// TIA Portal project "ESTHER_Gas_v4.0_4" (V13)

(* hardware
DEVICE "SIMATIC 1200 station_1"  S71200.Device
   slot 0: "S7-1200 rack"  Rack  V1.0
   slot 1: "PLC_1"  CPU 1215C DC/DC/DC  6ES7 215-1AG40-0XB0  V4.1
   slot 2: "DQ 16x24VDC_1"  6ES7 222-1BH32-0XB0  V2.0
   slot 3: "AI 8x13BIT_1"  6ES7 231-4HF32-0XB0  V2.0
   slot 4: "AI 8x13BIT_2"  6ES7 231-4HF32-0XB0  V2.0
   slot 101: "CM 1241 (RS422/485)_1"  6ES7 241-1CH32-0XB0  V2.1
   slot 102: "CM 1241 (RS422/485)_2"  6ES7 241-1CH32-0XB0  V2.1
*)

// ===== PLC "PLC_1"  CPU 1215C DC/DC/DC =====

VAR_GLOBAL   // PLC tag table "Default tag table"
   "PV701_NOT_CLOSED_LS" AT %I0.0 : Bool;   // PV701 Limit Switch
   "PV701_NOT_OPEN_LS" AT %I0.1 : Bool;   // PV701 Limit Switch
   "PV702_NOT_CLOSED_LS" AT %I0.2 : Bool;   // PV702 Limit Switch
   "PV702_NOT_OPEN_LS" AT %I0.3 : Bool;   // PV702 Limit Switch
   "PV703A_NOT_OPEN_LS" AT %I0.4 : Bool;
   "PV703A_NOT_CLOSED_LS" AT %I0.5 : Bool;
   "PV703B_NOT_OPEN_LS" AT %I0.6 : Bool;
   "PV703B_NOT_CLOSED_LS" AT %I0.7 : Bool;
   "PT101_ADC" AT %IW114 : Word;
   "PV101_NC" AT %Q9.3 : Bool;   // NC
   "PV102_NO" AT %Q9.4 : Bool;   // NO Temp
   "STEP_0_ON" AT %Q1.7 : Bool;
   "STEP_1_ON" AT %Q1.2 : Bool;
   "STEP_2_ON" AT %Q1.3 : Bool;
   "STEP_3_ON" AT %Q1.4 : Bool;
   "PV201_NC" AT %Q8.3 : Bool;
   "PV301_NC" AT %Q8.6 : Bool;
   "PV401_NC" AT %Q8.0 : Bool;
   "PV202_NC" AT %Q8.4 : Bool;   // NC Temp
   "PV302_NC" AT %Q8.7 : Bool;   // NC Temp
   "PV203_NO" AT %Q8.5 : Bool;   // NO Temp
   "PV303_NO" AT %Q0.3 : Bool;   // NO Temp
   "ABORT_ON" AT %Q1.5 : Bool;
   "START" AT %M0.0 : Bool;
   "STOP" AT %M0.1 : Bool;
   "PT502_VAL" AT %MD236 : Real;
   "DebugR" AT %MD184 : Real;
   "PT901_SP_O" AT %MD468 : Real;
   "PT901_SP_HE1" AT %MD472 : Real;
   "PT901_SP_HE2" AT %MD480 : Real;
   "PT901_SP_H" AT %MD476 : Real;
   "STEP_0_GO" AT %M2.0 : Bool;
   "PT901_SP_N" AT %MD484 : Real;
   "STEP_1_GO" AT %M2.1 : Bool;
   "ABORT_STOP" AT %M4.7 : Bool;
   "PT901_HIGH" AT %MD440 : Real;
   "STEP_2_GO" AT %M2.2 : Bool;
   "PT201_LOW" AT %MD404 : Real;
   "PT301_LOW" AT %MD408 : Real;
   "PT401_LOW" AT %MD412 : Real;
   "PT501_LOW" AT %MD416 : Real;
   "STEP_3_GO" AT %M2.3 : Bool;
   "STEP_4_GO" AT %M2.4 : Bool;
   "STEP_5_GO" AT %M2.5 : Bool;
   "STEP_6_GO" AT %M2.6 : Bool;
   "STEP_7_GO" AT %M2.7 : Bool;
   "STEP_4_ON" AT %M3.4 : Bool;
   "STEP_5_ON" AT %M3.5 : Bool;
   "STEP_6_ON" AT %M3.6 : Bool;
   "STEP_7_ON" AT %M3.7 : Bool;
   "PV501_NC" AT %Q9.5 : Bool;
   "PV402_NC" AT %Q8.1 : Bool;   // NC Temp
   "PV502_NC" AT %Q9.6 : Bool;   // NC Temp
   "PV601_NC" AT %Q9.0 : Bool;   // NC Temp
   "PV602_NC" AT %Q9.1 : Bool;   // NC Temp
   "PV603_NC" AT %Q9.2 : Bool;   // NC Temp
   "PV403_NO" AT %Q8.2 : Bool;   // NO Temp
   "PV503_NO" AT %Q9.7 : Bool;   // NO Temp
   "PV701_NC" AT %Q0.4 : Bool;   // NC With LS Temp
   "PV702_NC" AT %Q0.5 : Bool;   // NC With LS Temp
   "PV703A_NO" AT %Q0.6 : Bool;
   "PV703B_NO" AT %Q0.7 : Bool;
   "PT102_VAL" AT %MD204 : Real;
   "PT202_VAL" AT %MD212 : Real;
   "PT302_VAL" AT %MD220 : Real;
   "PT801_VAL" AT %MD244 : Real;
   "PT402_VAL" AT %MD228 : Real;
   "PT101_VAL" AT %MD200 : Real;
   "PT201_VAL" AT %MD208 : Real;
   "Clock_Byte" AT %MB100 : Byte;
   "Clock_2.5Hz" AT %M100.2 : Bool;
   "Clock_2Hz" AT %M100.3 : Bool;
   "Clock_1.25Hz" AT %M100.4 : Bool;
   "Clock_1Hz" AT %M100.5 : Bool;
   "Clock_0.625Hz" AT %M100.6 : Bool;
   "Clock_0.5Hz" AT %M100.7 : Bool;
   "System_Byte" AT %MB1 : Byte;
   "FirstScan" AT %M1.0 : Bool;
   "DiagStatusUpdate" AT %M1.1 : Bool;
   "AlwaysTRUE" AT %M1.2 : Bool;
   "AlwaysFALSE" AT %M1.3 : Bool;
   "STEP_9_ON" AT %M4.0 : Bool;
   "STEP_1_M" AT %M4.1 : Bool;
   "STEP_2_M" AT %M4.2 : Bool;
   "PT102_HIGH" AT %MD444 : Real;
   "PT202_HIGH" AT %MD448 : Real;
   "PT302_HIGH" AT %MD452 : Real;
   "PT402_HIGH" AT %MD456 : Real;
   "PT502_HIGH" AT %MD460 : Real;
   "PT601_HIGH" AT %MD464 : Real;
   "PT501_VAL" AT %MD232 : Real;
   "PT301_VAL" AT %MD216 : Real;
   "PT401_VAL" AT %MD224 : Real;
   "PT601_VAL" AT %MD240 : Real;
   "PT901_VAL" AT %MD248 : Real;
   "S0_0" AT %M101.0 : Bool;
   "S0_1" AT %M101.1 : Bool;
   "S0_END" AT %M101.7 : Bool;
   "S1_0" AT %M102.0 : Bool;
   "S1_1" AT %M102.1 : Bool;
   "S1_2" AT %M102.2 : Bool;
   "S1_3" AT %M102.3 : Bool;
   "S1_4" AT %M102.4 : Bool;
   "S1_5" AT %M102.5 : Bool;
   "S1_6" AT %M102.6 : Bool;
   "S1_7" AT %M102.7 : Bool;
   "S1_8" AT %M103.0 : Bool;
   "S1_9" AT %M103.1 : Bool;
   "S1_10" AT %M103.2 : Bool;
   "S1_11" AT %M103.3 : Bool;
   "S1_12" AT %M103.4 : Bool;
   "S1_13" AT %M103.5 : Bool;
   "ALARM" AT %M0.2 : Bool;
   "ALARM_CLR" AT %M0.3 : Bool;
   "PT102_CALC_90PRCT" AT %MD280 : Real;
   "S1_END" AT %M103.7 : Bool;
   "ALARM_PT101" AT %M20.0 : Bool;
   "ALARM_PT102" AT %M20.1 : Bool;
   "ALARM_PT201" AT %M20.2 : Bool;
   "ALARM_PT202" AT %M20.3 : Bool;
   "ALARM_PT301" AT %M20.4 : Bool;
   "ALARM_PT302" AT %M20.5 : Bool;
   "ALARM_PT401" AT %M20.6 : Bool;
   "ALARM_PT402" AT %M20.7 : Bool;
   "ALARM_PT501" AT %M21.0 : Bool;
   "ALARM_PT502" AT %M21.1 : Bool;
   "ALARM_PT601" AT %M21.2 : Bool;
   "ALARM_PT801" AT %M21.3 : Bool;
   "ALARM_PT901" AT %M21.4 : Bool;
   "TempReal_A" AT %MD188 : Real;
   "TempReal_B" AT %MD192 : Real;
   "TempWord_B" AT %MW144 : Word;
   "TempDWord_A" AT %MD160 : DInt;
   "TempWord_A" AT %MW140 : Word;
   "TempDWord_B" AT %MD164 : DInt;
   "LOOP_SEVEN_OK_S1" AT %M130.0 : Bool;
   "S1_14" AT %M103.6 : Bool;
   "ABORT_START" AT %M4.3 : Bool;
   "SA_0" AT %M116.0 : Bool;
   "SA_1" AT %M116.1 : Bool;
   "SA_END" AT %M116.7 : Bool;
   "SA_2" AT %M116.2 : Bool;
   "SA_M" AT %M116.6 : Bool;
   "S2_0" AT %M104.0 : Bool;
   "S2_1" AT %M104.1 : Bool;
   "S2_2" AT %M104.2 : Bool;
   "S2_3" AT %M104.3 : Bool;
   "S2_4" AT %M104.4 : Bool;
   "S2_5" AT %M104.5 : Bool;
   "S2_6" AT %M104.6 : Bool;
   "S2_7" AT %M104.7 : Bool;
   "PT202_CALC_10PRCT" AT %MD284 : Real;
   "S2_END" AT %M105.7 : Bool;
   "S3_0" AT %M106.0 : Bool;
   "S3_1" AT %M106.1 : Bool;
   "S3_2" AT %M106.2 : Bool;
   "S3_3" AT %M106.3 : Bool;
   "S3_4" AT %M106.4 : Bool;
   "S3_5" AT %M106.5 : Bool;
   "S3_6" AT %M106.6 : Bool;
   "S3_7" AT %M106.7 : Bool;
   "S3_END" AT %M107.7 : Bool;
   "MFC201_FLOW_MEAS" AT %MW256 : UInt;   // MFC Measure, Range 0....(32000)...41942
   "MFC401_FLOW_MEAS" AT %MW264 : UInt;   // MFC Measure, Range 0....(32000)...41942
   "MFC601_FLOW_MEAS" AT %MW272 : UInt;
   "AUTO_CYCLE" AT %M0.4 : Bool;
   "S0_M" AT %M101.3 : Bool;
   "MFC201_VOL_MEAS" AT %MW260 : UInt;
   "MFC401_VOL_MEAS" AT %MW268 : UInt;
   "MFC601_VOL_MEAS" AT %MW276 : UInt;
   "MFC201_FLOW_MAX" AT %MW258 : UInt;   // MFC User SetPoint, Range 0....32000
   "MFC401_FLOW_MAX" AT %MW266 : UInt;
   "S3_8" AT %M107.0 : Bool;
   "S3_9" AT %M107.1 : Bool;
   "S3_10" AT %M107.2 : Bool;
   "S3_11" AT %M107.3 : Bool;
   "PT302_CALC_90PRCT" AT %MD288 : Real;
   "S1_M" AT %M101.4 : Bool;
   "S2_M" AT %M105.0 : Bool;
   "S3_M" AT %M107.4 : Bool;
   "S4_0" AT %M108.0 : Bool;
   "S4_1" AT %M108.1 : Bool;
   "S4_2" AT %M108.2 : Bool;
   "S4_3" AT %M108.3 : Bool;
   "S4_4" AT %M108.4 : Bool;
   "S4_5" AT %M108.5 : Bool;
   "S4_END" AT %M109.7 : Bool;
   "S4_M" AT %M109.6 : Bool;
   "S4_6" AT %M108.6 : Bool;
   "S4_7" AT %M108.7 : Bool;
   "S4_8" AT %M109.0 : Bool;
   "S4_9" AT %M109.1 : Bool;
   "S4_10" AT %M109.2 : Bool;
   "TEST_START" AT %M0.5 : Bool;
   "TEST_STOP" AT %M0.6 : Bool;
   "TEST_ON" AT %M0.7 : Bool;
   "ST_END" AT %M120.7 : Bool;
   "ST_0" AT %M117.0 : Bool;
   "ST_1" AT %M117.1 : Bool;
   "TEST_GO" AT %M3.0 : Bool;
   "ST_2" AT %M117.2 : Bool;
   "ST_3" AT %M117.3 : Bool;
   "ST_4" AT %M117.4 : Bool;
   "ST_5" AT %M117.5 : Bool;
   "PT801_SAVE" AT %MD324 : Real;
   "S5_END" AT %M111.7 : Bool;
   "S5_0" AT %M110.0 : Bool;
   "S5_1" AT %M110.1 : Bool;
   "S5_2" AT %M110.2 : Bool;
   "S5_3" AT %M110.3 : Bool;
   "S5_4" AT %M110.4 : Bool;
   "S5_M" AT %M111.6 : Bool;
   "PT502_CALC_90PRCT" AT %MD296 : Real;
   "S5_5" AT %M110.5 : Bool;
   "S5_6" AT %M110.6 : Bool;
   "S5_7" AT %M110.7 : Bool;
   "S5_8" AT %M111.0 : Bool;
   "ST_6" AT %M117.6 : Bool;
   "ST_7" AT %M117.7 : Bool;
   "ST_8" AT %M118.0 : Bool;
   "ST_M" AT %M120.6 : Bool;
   "ST_9" AT %M118.1 : Bool;
   "ST_10" AT %M118.2 : Bool;
   "ST_11" AT %M118.3 : Bool;
   "ST_12" AT %M118.4 : Bool;
   "ST_13" AT %M118.5 : Bool;
   "ST_14" AT %M118.6 : Bool;
   "ST_15" AT %M118.7 : Bool;
   "TEST_FAIL" AT %M3.1 : Bool;
   "ST_16" AT %M119.0 : Bool;
   "ST_17" AT %M119.1 : Bool;
   "ST_18" AT %M119.2 : Bool;
   "ST_19" AT %M119.3 : Bool;
   "PT301_SAVE" AT %MD316 : Real;
   "PT501_SAVE" AT %MD320 : Real;
   "ST_20" AT %M119.4 : Bool;
   "ST_21" AT %M119.5 : Bool;
   "ST_22" AT %M119.6 : Bool;
   "PT101_SAVE" AT %MD312 : Real;
   "ST_23" AT %M119.7 : Bool;
   "S6_0" AT %M112.0 : Bool;
   "S6_1" AT %M112.1 : Bool;
   "S6_END" AT %M113.7 : Bool;
   "S6_M" AT %M113.6 : Bool;
   "S6_2" AT %M112.2 : Bool;
   "S6_3" AT %M112.3 : Bool;
   "S6_4" AT %M112.4 : Bool;
   "S6_5" AT %M112.5 : Bool;
   "PT401_CALC_50PRCT" AT %MD328 : Real;
   "S6_6" AT %M112.6 : Bool;
   "S6_7" AT %M112.7 : Bool;
   "S6_8" AT %M113.0 : Bool;
   "S6_9" AT %M113.1 : Bool;
   "PT102_ADC" AT %IW112 : Word;
   "STEP_9_GO" AT %M3.2 : Bool;
   "Tag_MB_MS" AT %M3.3 : Bool;
   "MB_MS_Done" AT %M4.4 : Bool;
   "MB_MS_Error" AT %M4.5 : Bool;
   "MB_MS_Status" AT %MW6 : Word;
   "MB_MST_CM_Done" AT %M4.6 : Bool;
   "MB_MST_CM_Error" AT %M5.0 : Bool;
   "MB_MST_CM_Status" AT %MW8 : Word;
   "S7_0" AT %M114.0 : Bool;
   "S7_1" AT %M114.1 : Bool;
   "S7_2" AT %M114.2 : Bool;
   "S7_3" AT %M114.3 : Bool;
   "S7_4" AT %M114.4 : Bool;
   "S7_5" AT %M114.5 : Bool;
   "S7_END" AT %M115.7 : Bool;
   "S7_M" AT %M115.6 : Bool;
   "S7_6" AT %M114.6 : Bool;
   "S7_7" AT %M114.7 : Bool;
   "S7_8" AT %M115.0 : Bool;
   "S7_9" AT %M115.1 : Bool;
   "S7_10" AT %M115.2 : Bool;
   "S7_11" AT %M115.3 : Bool;
   "S7_12" AT %M115.4 : Bool;
   "MB_SLV_CM_Done" AT %M5.1 : Bool;
   "MB_SLV_CM_Error" AT %M5.2 : Bool;
   "MB_SLV_CM_Status" AT %MW14 : Word;
   "MB_SLV_Error" AT %M5.3 : Bool;
   "MB_SLV_Status" AT %MW16 : Word;
   "PT101_Norm" AT %MD340 : Real;
   "PT101_LOW" AT %MD392 : Real;
   "PT201_ADC" AT %IW122 : Word;
   "PT202_ADC" AT %IW120 : Word;
   "PT301_ADC" AT %IW126 : Word;
   "PT302_ADC" AT %IW124 : Word;
   "PT501_ADC" AT %IW118 : Word;
   "PT801_ADC" AT %IW136 : Word;
   "PT502_ADC" AT %IW116 : Word;
   "PT102_Norm" AT %MD344 : Real;
   "PT201_Norm" AT %MD348 : Real;
   "PT202_Norm" AT %MD352 : Real;
   "PT301_Norm" AT %MD356 : Real;
   "PT302_Norm" AT %MD360 : Real;
   "PT501_Norm" AT %MD364 : Real;
   "PT502_Norm" AT %MD368 : Real;
   "PT801_Norm" AT %MD372 : Real;
   "PT401_Norm" AT %MD376 : Real;
   "PT402_Norm" AT %MD380 : Real;
   "PT601_Norm" AT %MD384 : Real;
   "PT901_Norm" AT %MD388 : Real;
   "S1_1A" AT %M65.0 : Bool;
   "PV70x_LS_FTS_TIME" AT %MD520 : Time;
   "PV70x_LS_WAIT_TIME" AT %MD524 : Time;
   "PV70x_LS_WAIT" AT %MD528 : Time;
   "ALARM_PV701_NOT_CLS" AT %M21.5 : Bool;
   "ALARM_PV701_NOT_OPN" AT %M21.6 : Bool;
   "ALARM_PV702_NOT_CLS" AT %M21.7 : Bool;
   "ALARM_PV702_NOT_OPN" AT %M22.0 : Bool;
   "ALARM_PV703A_NOT_CLS" AT %M22.1 : Bool;
   "ALARM_PV703A_NOT_OPN" AT %M22.2 : Bool;
   "ALARM_PV703B_NOT_CLS" AT %M22.3 : Bool;
   "ALARM_PV703B_NOT_OPN" AT %M22.4 : Bool;
   "S1_10A" AT %M65.1 : Bool;
   "tempLS1" AT %M5.4 : Bool;
   "tempLS2" AT %M5.5 : Bool;
   "ALARM_BREAKPOINT" AT %M22.5 : Bool;
   "S2_4A" AT %M65.4 : Bool;
   "S3_4A" AT %M65.5 : Bool;
   "S3_5A" AT %M65.6 : Bool;
   "S3_7A" AT %M65.7 : Bool;
   "S3_8A" AT %M66.0 : Bool;
   "ST_1A" AT %M70.0 : Bool;
   "ST_24" AT %M120.0 : Bool;
   "TEST_PV0" AT %M30.0 : Bool;
   "TEST_PV1" AT %M30.1 : Bool;
   "TEST_PV2" AT %M30.2 : Bool;
   "TEST_PV3" AT %M30.3 : Bool;
   "PT401_ADC" AT %IW134 : Word;
   "PT901_ADC" AT %IW130 : Word;
   "PT601_ADC" AT %IW128 : Word;
   "PT402_ADC" AT %IW132 : Word;
   "PT801_99" AT %MD332 : Real;
   "temp702_LS_ET" AT %MD10 : Time;
   "temp702_LS_Count" AT %MD24 : Time;
   "Tag_MB_EN" AT %M5.6 : Bool;
   "Tag_MB_REQ" AT %M5.7 : Bool;
   "MB_MS_Busy" AT %M18.0 : Bool;
   "MS_MS_DONE_LED" AT %M18.1 : Bool;
   "TEMP_MFC_SAVE" AT %MW602 : Word;
   "Tag_MB_CLR" AT %M18.2 : Bool;
   "PULSE_NUMBER" AT %MW28 : UInt;
   "MB_MS_STATUS_SAV" AT %MW606 : Word;
   "Clock_5Hz" AT %M100.1 : Bool;
   "Clock_10Hz" AT %M100.0 : Bool;
   "MFC_FLOW_NORM" AT %MD600 : Real;
   "MFC601_FLOW_MAX" AT %MW274 : UInt;
   "SA_3" AT %M116.3 : Bool;
   "SA_4" AT %M116.4 : Bool;
   "SA_5" AT %M116.5 : Bool;
   "PT901_SAVE" AT %MD336 : Real;
   "S1_7A" AT %M65.2 : Bool;
   "SMB_0" AT %M121.0 : Bool;
   "SMB_END" AT %M122.7 : Bool;
   "SMB_1" AT %M121.1 : Bool;
   "SMB_2" AT %M121.2 : Bool;
   "SMB_3" AT %M121.3 : Bool;
   "SMB_4" AT %M121.4 : Bool;
   "SMB_5" AT %M121.5 : Bool;
   "SMB_6" AT %M121.6 : Bool;
   "SMB_7" AT %M121.7 : Bool;
   "SMB_8" AT %M122.0 : Bool;
   "SMB_M" AT %M122.6 : Bool;
   "S4_5A" AT %M109.3 : Bool;
   "S4_8A" AT %M109.4 : Bool;
   "S9_0" AT %M123.0 : Bool;
   "S9_1" AT %M123.1 : Bool;
   "S9_2" AT %M123.2 : Bool;
   "S9_END" AT %M124.7 : Bool;
   "S9_3" AT %M123.3 : Bool;
   "S9_4" AT %M123.4 : Bool;
   "S6_3A" AT %M113.2 : Bool;
   "MFC401_VOL_SP" AT %MW626 : UInt;
   "SMB_9" AT %M122.1 : Bool;
   "S7_5A" AT %M115.5 : Bool;
   "S1_10B" AT %M65.3 : Bool;
   "S9_1A" AT %M123.5 : Bool;
   "S9_2A" AT %M123.6 : Bool;
   "TimerS1_1_wait" AT %MD80 : Time;
   "TimerS1_2_wait" AT %MD84 : Time;
   "S9_M" AT %M124.6 : Bool;
   "S7_0A" AT %M120.1 : Bool;
   "TimerS1_3_wait" AT %MD88 : Time;
   "TimerTests_1_wait" AT %MD92 : Time;
   "PT901_SP_N_ZERO" AT %MD488 : Real;
   "TimerS9_1_wait" AT %MD96 : Time;
   "MFC601_VOL_HE1_SAVE" AT %MW632 : UInt;
   "MFC601_VOL_HE2_SAVE" AT %MW634 : UInt;
   "PT901_END_O" AT %MD496 : Real;
   "PT901_END_HE1" AT %MD500 : Real;
   "PT901_END_H" AT %MD504 : Real;
   "PT901_END_HE2" AT %MD508 : Real;
   "PT901_END_S1" AT %MD492 : Real;
   "ABORT_BUTTON" AT %I1.0 : Bool;
   "SMB_10" AT %M122.2 : Bool;
   "Counter_S1" AT %MW78 : UInt;
   "S7_1A" AT %M120.2 : Bool;
   "TimerS1_left" AT %MD636 : Time;
   "MFC201_VOL_FMEAS" AT %MD610 : Real;
   "MFC401_VOL_FMEAS" AT %MD614 : Real;
   "MFC601_VOL_FMEAS" AT %MD618 : Real;
   "MFC201_FLOW_FMEAS" AT %MD640 : Real;
   "MFC401_FLOW_FMEAS" AT %MD644 : Real;
   "MFC601_FLOW_FMEAS" AT %MD648 : Real;
   "S4_5B" AT %M109.5 : Bool;
   "S7_2A" AT %M120.3 : Bool;
   "S6_3B" AT %M113.3 : Bool;
   "S6_3C" AT %M113.4 : Bool;
   "S7_1B" AT %M120.4 : Bool;
   "S4_2A" AT %M107.5 : Bool;
   "MFC201_FTEMP" AT %MD652 : Real;
   "MFC401_FTEMP" AT %MD656 : Real;
   "MFC601_FTEMP" AT %MD660 : Real;
   "PT901_RAW" AT %MD684 : Real;
   "PT601_RAW" AT %MD680 : Real;
   "ON" AT %Q1.6 : Bool;
   "RED_LIGHT" AT %Q0.0 : Bool;
   "YELLOW_LIGHT" AT %Q0.1 : Bool;
   "GREEN_LIGHT" AT %Q0.2 : Bool;
   "DOORS_LOCK" AT %Q1.1 : Bool;
   "BUZZER" AT %Q1.0 : Bool;
   "BUZZER_ON" AT %M130.1 : Bool;
   "RED_ON" AT %M130.2 : Bool;
   "RED_BLINK" AT %M130.3 : Bool;
   "DOORS_CLOSED" AT %I1.1 : Bool;
   "ALARM_DOORS_OPEN" AT %M22.6 : Bool;
   "PT801_LOW" AT %MD420 : Real;
END_VAR

VAR_GLOBAL CONSTANT   // PLC tag table "Default tag table"
   "MB_AD_OPERATION" : UDInt := 40032;
   "MB_AD_WINK" : UDInt := 40001;
   "MB_AD_SETPOINT" : UDInt := 40034;
   "MB_AD_TEMPERATURE" : UDInt := 41064;
   "MB_AD_ALARM" : UDInt := 43106;
   "MB_AD_COUNTER_VAL" : UDInt := 43330;
   "MB_AD_COUNTER_LIMIT" : UDInt := 43332;
   "MB_AD_COUNTER_SP_MODE" : UDInt := 43334;
   "MB_AD_COUNTER_NEW_SP" : UDInt := 43335;
   "MB_AD_CONTROL_MODE" : UDInt := 40037;
   "MB_AD_ALARM_SP_MODE" : UDInt := 43110;
   "MB_VAL_WINK" : UInt := 0;
   "MB_VAL_CONTROL_MODE_BUS" : UInt := 0;
   "MB_VAL_CONTROL_MODE_CLOSE" : UInt := 3;
   "MB_VAL_CONTROL_MODE_SP_100" : UInt := 7;
   "MB_VAL_CONTROL_MODE_OPEN" : UInt := 8;
   "MB_VAL_CONTROL_MODE_SP_0" : UInt := 12;
   "MB_VAL_COUNT_MODE_OFF" : UInt := 0;
   "MB_VAL_COUNT_MODE_UP" : UInt := 1;
   "MB_VAL_COUNT_MODE_UP_LIMIT" : UInt := 2;
   "MB_VAL_COUNT_SP_MODE_NO_CHANGE" : UInt := 0;
   "MB_VAL_COUNT_SP_MODE_CHANGE" : UInt := 1;
   "MB_AD_COUNTER_MODE" : UDInt := 43337;
   "MB_AD_COUNTER_RST_ENABL" : UDInt := 43338;
   "MB_VAL_COUNT_RST_ENABL" : UInt := 5;
   "MB_AD_RESET" : UDInt := 43689;
   "MB_VAL_RST_COUNTER" : UInt := 3;   // Send 0 first
   "MB_VAL_RST_SOFT" : UInt := 5;
   "MFC_201_MB_ADDR" : USInt := 20;
   "MFC_401_MB_ADDR" : USInt := 40;
   "MFC_601_MB_ADDR" : USInt := 60;
   "MFC_201_CAPACITY" : Real := 2.0;
   "MFC_401_CAPACITY" : Real := 5.95;
   "MFC_601_CAPACITY" : Real := 50.0;
   "MFC_FLOW_100_W" : UInt := 32000;
   "MFC_FLOW_50_W" : UInt := 16000;
   "MFC_401_INIT_MAX_FLOW" : UInt := 2700;
   "MFC_201_INIT_MAX_FLOW" : UInt := 3200;
   "MB_AD_COUNTER_UNIT_IDX" : UDInt := 43331;
   "MB_VAL_COUNT_UNIT_IDX_mLn" : UInt := 2;   // mln
   "PT302_ZERO" : Real := 1.4;   // System clogged. Should be 0.2
   "PT202_ZERO" : Real := 1.8;   // System clogged. Should be 0.3
   "PT601_ZERO" : Real := 1.2;   // System clogged
   "PT901_SP_PV703B_OPEN" : Real := 2.0;
   "PT901_ZERO" : Real := 0.0;
   "PT801_LOW_C" : Real := 20.0;
   "PT101_LOW_C" : Real := 110.0;
   "PT502_ZERO" : Real := 0.9;   // System clogged. Should be -0.5
   "PT201_ZERO" : Real := -1.0;
   "PT901_HIGH_N" : Real := 10.0;
   "PT901_HIGH_O" : Real := 12.6;
   "PT901_HIGH_HE1" : Real := 80.1;
   "PT901_HIGH_H" : Real := 99.6;
   "PT901_HIGH_HE2" : Real := 100.1;
   "PT901_HIGH_PV703B" : Real := 10.0;
   "PT901_DELTA" : Real := 4.0;
   "PT301_LOW_C" : Real := 140.0;
   "PT501_LOW_C" : Real := -10.0;
   "PT201_LOW_C" : Real := 35.0;
   "PT401_LOW_C" : Real := 137.0;
   "PT202_ZERO_MAX" : Real := 0.6;
   "PT102_ZERO_1" : Real := 0.2;
   "MB_AD_COUNTER_UNIT_INDEX" : UDInt := 43331;
   "MB_AD_TEMP_FLOAT" : UDInt := 441273;
   "MB_AD_COUNTER_LIMIT_FLOAT" : UDInt := 459417;
   "PT901_OFFSET" : Real := -0.17;
   "PT601_OFFSET" : Real := 1.0;
   "STEP1_LOOPS" : UInt := 3;
   "STEP1_MFC_FL_SP" : UInt := 30000;
   "MB_MODE_READ" : UInt := 0;
   "MB_MODE_WRITE" : UInt := 1;
   "PT502_HIGH_C" : Real := 120.0;
   "PT302_HIGH_C" : Real := 120.0;
END_VAR

TYPE "UDT_DATA_PTR"
VERSION : 0.1
   STRUCT
      DATA : Array[0..6] of Int;
   END_STRUCT;
END_TYPE

TYPE "UDT_DATA_REAL_PTR"
   STRUCT
      DATA : Array[0..1] of Real;
   END_STRUCT;
END_TYPE

DATA_BLOCK "MB_DATA_MFC"   // DB23
{ S7_Optimized_Access := 'FALSE' }
VERSION : 0.1
   VAR
      OPERATION : Struct
      END_STRUCT;
      TEMPERATURE : UInt;
      ALARM : Struct
      END_STRUCT;
      "COUNTER" : Struct
      END_STRUCT;
      PARAM : Struct
      END_STRUCT;
      "STEP" : UInt;
      MB_WRT_PARAM : Struct
      END_STRUCT;
      MB_MASTER_ENABLE : Bool;
      MB_WRT_FLAG : Bool;
      MB_WRT_FLAG_SAVE : Bool;
   END_VAR
BEGIN
END_DATA_BLOCK

DATA_BLOCK "MB_DATA_MX"   // DB42
{ S7_Optimized_Access := 'FALSE' }
VERSION : 0.1
   VAR
      MEASURE : Struct
      END_STRUCT;
      ALARM_STATUS : Struct
      END_STRUCT;
      SEC_COUNTER : UInt;
      PARAM : Struct
      END_STRUCT;
      "STEP" : UInt;
      MB_WRT_PARAM : Struct
      END_STRUCT;
      MB_MASTER_ENABLE : Bool;
      MB_WRT_FLAG : Bool;
      MB_WRT_FLAG_SAVE : Bool;
      MS_Status : Word;
      MS_Done : Bool;
      MS_Busy : Bool;
      MS_Error : Bool;
      MS_Clock_tag : Bool;
      MS_Status_Save : Word;
   END_VAR
BEGIN
END_DATA_BLOCK

DATA_BLOCK "MB_MFC_FLOAT_DB"   // DB47
{ S7_Optimized_Access := 'FALSE' }
VERSION : 0.1
// stored: InstanceOfName MB_MFC_FLOAT
"MB_MFC_FLOAT"
BEGIN
END_DATA_BLOCK

DATA_BLOCK "MB_MFC_INT_DB"   // DB51
{ S7_Optimized_Access := 'FALSE' }
VERSION : 0.1
// stored: InstanceOfName MB_MFC_INT
"MB_MFC_INT"
BEGIN
END_DATA_BLOCK

// folder: System blocks/Program resources

DATA_BLOCK "IEC_Timer_S1_DB5"   // DB1
{ S7_Optimized_Access := 'FALSE' }
AUTHOR : Simatic
FAMILY : IEC
NAME : IEC_TMR
VERSION : 1.0
// stored: InstanceOfName ?
"?"
BEGIN
END_DATA_BLOCK

DATA_BLOCK "IEC_Timer_ALM_PV703B_CLS_DB"   // DB2
{ S7_Optimized_Access := 'FALSE' }
AUTHOR : Simatic
FAMILY : IEC
NAME : IEC_TMR
VERSION : 1.0
// stored: InstanceOfName ?
"?"
BEGIN
END_DATA_BLOCK

DATA_BLOCK "IEC_Timer_S1_DB3"   // DB3
{ S7_Optimized_Access := 'FALSE' }
AUTHOR : Simatic
FAMILY : IEC
NAME : IEC_TMR
VERSION : 1.0
// stored: InstanceOfName ?
"?"
BEGIN
END_DATA_BLOCK

DATA_BLOCK "Timer_S1_DB_1S"   // DB4
{ S7_Optimized_Access := 'FALSE' }
AUTHOR : Simatic
FAMILY : IEC
NAME : IEC_TMR
VERSION : 1.0
// stored: InstanceOfName ?
"?"
BEGIN
END_DATA_BLOCK

DATA_BLOCK "Timer_S3_DB_1S"   // DB5
{ S7_Optimized_Access := 'FALSE' }
AUTHOR : Simatic
FAMILY : IEC
NAME : IEC_TMR
VERSION : 1.0
// stored: InstanceOfName ?
"?"
BEGIN
END_DATA_BLOCK

DATA_BLOCK "IEC_Counter_S1_1"   // DB6
{ S7_Optimized_Access := 'FALSE' }
AUTHOR : Simatic
FAMILY : IEC
NAME : UCNTR
VERSION : 1.2
// stored: InstanceOfName ?
"?"
BEGIN
END_DATA_BLOCK

DATA_BLOCK "IEC_Timer_0_DB_1"   // DB7
{ S7_Optimized_Access := 'FALSE' }
AUTHOR : Simatic
FAMILY : IEC
NAME : IEC_TMR
VERSION : 1.0
// stored: InstanceOfName ?
"?"
BEGIN
END_DATA_BLOCK

DATA_BLOCK "IEC_Counter_MB_DB"   // DB8
{ S7_Optimized_Access := 'FALSE' }
AUTHOR : Simatic
FAMILY : IEC
NAME : UCNTR
VERSION : 1.2
// stored: InstanceOfName ?
"?"
BEGIN
END_DATA_BLOCK

DATA_BLOCK "IEC_Counter_MXT_DB"   // DB9
{ S7_Optimized_Access := 'FALSE' }
AUTHOR : Simatic
FAMILY : IEC
NAME : UCNTR
VERSION : 1.2
// stored: InstanceOfName ?
"?"
BEGIN
END_DATA_BLOCK

DATA_BLOCK "IEC_Timer_S2_1"   // DB10
{ S7_Optimized_Access := 'FALSE' }
AUTHOR : Simatic
FAMILY : IEC
NAME : IEC_TMR
VERSION : 1.0
// stored: InstanceOfName ?
"?"
BEGIN
END_DATA_BLOCK

DATA_BLOCK "IEC_Timer_S2_2"   // DB11
{ S7_Optimized_Access := 'FALSE' }
AUTHOR : Simatic
FAMILY : IEC
NAME : IEC_TMR
VERSION : 1.0
// stored: InstanceOfName ?
"?"
BEGIN
END_DATA_BLOCK

DATA_BLOCK "IEC_Timer_1_ST1_DB"   // DB12
{ S7_Optimized_Access := 'FALSE' }
AUTHOR : Simatic
FAMILY : IEC
NAME : IEC_TMR
VERSION : 1.0
// stored: InstanceOfName ?
"?"
BEGIN
END_DATA_BLOCK

DATA_BLOCK "IEC_Timer_T2_1s_DB"   // DB13
{ S7_Optimized_Access := 'FALSE' }
AUTHOR : Simatic
FAMILY : IEC
NAME : IEC_TMR
VERSION : 1.0
// stored: InstanceOfName ?
"?"
BEGIN
END_DATA_BLOCK

DATA_BLOCK "Timer_S4_DB_1S"   // DB14
{ S7_Optimized_Access := 'FALSE' }
AUTHOR : Simatic
FAMILY : IEC
NAME : IEC_TMR
VERSION : 1.0
// stored: InstanceOfName ?
"?"
BEGIN
END_DATA_BLOCK

DATA_BLOCK "IEC_Timer_T2_2_DB"   // DB15
{ S7_Optimized_Access := 'FALSE' }
AUTHOR : Simatic
FAMILY : IEC
NAME : IEC_TMR
VERSION : 1.0
// stored: InstanceOfName ?
"?"
BEGIN
END_DATA_BLOCK

DATA_BLOCK "IEC_Timer_ST_DB_1"   // DB16
{ S7_Optimized_Access := 'FALSE' }
AUTHOR : Simatic
FAMILY : IEC
NAME : IEC_TMR
VERSION : 1.0
// stored: InstanceOfName ?
"?"
BEGIN
END_DATA_BLOCK

DATA_BLOCK "IEC_Timer_S5_DB_1"   // DB17
{ S7_Optimized_Access := 'FALSE' }
AUTHOR : Simatic
FAMILY : IEC
NAME : IEC_TMR
VERSION : 1.0
// stored: InstanceOfName ?
"?"
BEGIN
END_DATA_BLOCK

DATA_BLOCK "IEC_Timer_S5_DB_2"   // DB18
{ S7_Optimized_Access := 'FALSE' }
AUTHOR : Simatic
FAMILY : IEC
NAME : IEC_TMR
VERSION : 1.0
// stored: InstanceOfName ?
"?"
BEGIN
END_DATA_BLOCK

DATA_BLOCK "IEC_Timer_S6_DB_1"   // DB19
{ S7_Optimized_Access := 'FALSE' }
AUTHOR : Simatic
FAMILY : IEC
NAME : IEC_TMR
VERSION : 1.0
// stored: InstanceOfName ?
"?"
BEGIN
END_DATA_BLOCK

DATA_BLOCK "IEC_Timer_MFC_RST_ODD_DB"   // DB20
{ S7_Optimized_Access := 'FALSE' }
AUTHOR : Simatic
FAMILY : IEC
NAME : IEC_TMR
VERSION : 1.0
// stored: InstanceOfName ?
"?"
BEGIN
END_DATA_BLOCK

DATA_BLOCK "IEC_Timer_S7_1A_DB"   // DB24
{ S7_Optimized_Access := 'FALSE' }
AUTHOR : Simatic
FAMILY : IEC
NAME : IEC_TMR
VERSION : 1.0
// stored: InstanceOfName ?
"?"
BEGIN
END_DATA_BLOCK

DATA_BLOCK "IEC_Timers_SMB_DB"   // DB25
{ S7_Optimized_Access := 'FALSE' }
AUTHOR : Simatic
FAMILY : IEC
NAME : IEC_TMR
VERSION : 1.0
// stored: InstanceOfName ?
"?"
BEGIN
END_DATA_BLOCK

DATA_BLOCK "IEC_Timer_MFC_RST_EVN_DB"   // DB26
{ S7_Optimized_Access := 'FALSE' }
AUTHOR : Simatic
FAMILY : IEC
NAME : IEC_TMR
VERSION : 1.0
// stored: InstanceOfName ?
"?"
BEGIN
END_DATA_BLOCK

DATA_BLOCK "IEC_Timer_MFC_WRT_EVEN_DB"   // DB27
{ S7_Optimized_Access := 'FALSE' }
AUTHOR : Simatic
FAMILY : IEC
NAME : IEC_TMR
VERSION : 1.0
// stored: InstanceOfName ?
"?"
BEGIN
END_DATA_BLOCK

DATA_BLOCK "IEC_Timer_ALM_PV701_CLS_DB"   // DB28
{ S7_Optimized_Access := 'FALSE' }
AUTHOR : Simatic
FAMILY : IEC
NAME : IEC_TMR
VERSION : 1.0
// stored: InstanceOfName ?
"?"
BEGIN
END_DATA_BLOCK

DATA_BLOCK "IEC_Timer_ALM_PV701_OPN_DB"   // DB29
{ S7_Optimized_Access := 'FALSE' }
AUTHOR : Simatic
FAMILY : IEC
NAME : IEC_TMR
VERSION : 1.0
// stored: InstanceOfName ?
"?"
BEGIN
END_DATA_BLOCK

DATA_BLOCK "IEC_Timer_ALM_PV702_CLS_DB"   // DB30
{ S7_Optimized_Access := 'FALSE' }
AUTHOR : Simatic
FAMILY : IEC
NAME : IEC_TMR
VERSION : 1.0
// stored: InstanceOfName ?
"?"
BEGIN
END_DATA_BLOCK

DATA_BLOCK "IEC_Timer_ALM_PV702_OPN_DB"   // DB31
{ S7_Optimized_Access := 'FALSE' }
AUTHOR : Simatic
FAMILY : IEC
NAME : IEC_TMR
VERSION : 1.0
// stored: InstanceOfName ?
"?"
BEGIN
END_DATA_BLOCK

DATA_BLOCK "IEC_Timer_ALM_PV703A_CLS_DB"   // DB32
{ S7_Optimized_Access := 'FALSE' }
AUTHOR : Simatic
FAMILY : IEC
NAME : IEC_TMR
VERSION : 1.0
// stored: InstanceOfName ?
"?"
BEGIN
END_DATA_BLOCK

DATA_BLOCK "IEC_Timer_ALM_PV703A_OPN_DB"   // DB33
{ S7_Optimized_Access := 'FALSE' }
AUTHOR : Simatic
FAMILY : IEC
NAME : IEC_TMR
VERSION : 1.0
// stored: InstanceOfName ?
"?"
BEGIN
END_DATA_BLOCK

DATA_BLOCK "IEC_Timer_ALM_PV703B_OPN_DB"   // DB34
{ S7_Optimized_Access := 'FALSE' }
AUTHOR : Simatic
FAMILY : IEC
NAME : IEC_TMR
VERSION : 1.0
// stored: InstanceOfName ?
"?"
BEGIN
END_DATA_BLOCK

DATA_BLOCK "IEC_Timer_WAIT_PV70x_DB"   // DB35
{ S7_Optimized_Access := 'FALSE' }
AUTHOR : Simatic
FAMILY : IEC
NAME : IEC_TMR
VERSION : 1.0
// stored: InstanceOfName ?
"?"
BEGIN
END_DATA_BLOCK

DATA_BLOCK "Timer_S1_DB_3S"   // DB36
{ S7_Optimized_Access := 'FALSE' }
AUTHOR : Simatic
FAMILY : IEC
NAME : IEC_TMR
VERSION : 1.0
// stored: InstanceOfName ?
"?"
BEGIN
END_DATA_BLOCK

DATA_BLOCK "Timer_S1_DB_5S"   // DB37
{ S7_Optimized_Access := 'FALSE' }
AUTHOR : Simatic
FAMILY : IEC
NAME : IEC_TMR
VERSION : 1.0
// stored: InstanceOfName ?
"?"
BEGIN
END_DATA_BLOCK

DATA_BLOCK "IEC_Timer_S1_DB4"   // DB38
{ S7_Optimized_Access := 'FALSE' }
AUTHOR : Simatic
FAMILY : IEC
NAME : IEC_TMR
VERSION : 1.0
// stored: InstanceOfName ?
"?"
BEGIN
END_DATA_BLOCK

DATA_BLOCK "IEC_Timer_S9_DB"   // DB39
{ S7_Optimized_Access := 'FALSE' }
AUTHOR : Simatic
FAMILY : IEC
NAME : IEC_TMR
VERSION : 1.0
// stored: InstanceOfName ?
"?"
BEGIN
END_DATA_BLOCK

DATA_BLOCK "IEC_Timer_S9_1_DB"   // DB40
{ S7_Optimized_Access := 'FALSE' }
AUTHOR : Simatic
FAMILY : IEC
NAME : IEC_TMR
VERSION : 1.0
// stored: InstanceOfName ?
"?"
BEGIN
END_DATA_BLOCK

DATA_BLOCK "IEC_Timer_S1_5m_DB3"   // DB41
{ S7_Optimized_Access := 'FALSE' }
AUTHOR : Simatic
FAMILY : IEC
NAME : IEC_TMR
VERSION : 1.0
// stored: InstanceOfName ?
"?"
BEGIN
END_DATA_BLOCK

DATA_BLOCK "IEC_Timer_Buzzer_DB"   // DB45
{ S7_Optimized_Access := 'FALSE' }
AUTHOR : Simatic
FAMILY : IEC
NAME : IEC_TMR
VERSION : 1.0
// stored: InstanceOfName ?
"?"
BEGIN
END_DATA_BLOCK

DATA_BLOCK "IEC_Timer_S4_2_DB"   // DB46
{ S7_Optimized_Access := 'FALSE' }
AUTHOR : Simatic
FAMILY : IEC
NAME : IEC_TMR
VERSION : 1.0
// stored: InstanceOfName ?
"?"
BEGIN
END_DATA_BLOCK

DATA_BLOCK "IEC_Timer_Buzzer_1_DB"   // DB49
{ S7_Optimized_Access := 'FALSE' }
AUTHOR : Simatic
FAMILY : IEC
NAME : IEC_TMR
VERSION : 1.0
// stored: InstanceOfName ?
"?"
BEGIN
END_DATA_BLOCK

DATA_BLOCK "IEC_Timer_S4_5B_DB"   // DB54
{ S7_Optimized_Access := 'FALSE' }
AUTHOR : Simatic
FAMILY : IEC
NAME : IEC_TMR
VERSION : 1.0
// stored: InstanceOfName ?
"?"
BEGIN
END_DATA_BLOCK

DATA_BLOCK "IEC_Timers_S7_0_DB"   // DB55
{ S7_Optimized_Access := 'FALSE' }
AUTHOR : Simatic
FAMILY : IEC
NAME : IEC_TMR
VERSION : 1.0
// stored: InstanceOfName ?
"?"
BEGIN
END_DATA_BLOCK

DATA_BLOCK "IEC_Timer_S7_1_DB"   // DB56
{ S7_Optimized_Access := 'FALSE' }
AUTHOR : Simatic
FAMILY : IEC
NAME : IEC_TMR
VERSION : 1.0
// stored: InstanceOfName ?
"?"
BEGIN
END_DATA_BLOCK

DATA_BLOCK "IEC_Timer_S7_2_DB"   // DB58
{ S7_Optimized_Access := 'FALSE' }
AUTHOR : Simatic
FAMILY : IEC
NAME : IEC_TMR
VERSION : 1.0
// stored: InstanceOfName ?
"?"
BEGIN
END_DATA_BLOCK

// folder: (top level)

FUNCTION_BLOCK "MB_MFC_FLOAT"   // FB1, LAD
{ S7_Optimized_Access := 'FALSE' }
VERSION : 0.1
// Step  -1: Stopped 
// Steps 0-4: measure float vals
// Step 10 : load FSetpoint
// Steps 20 : load Counter Limit  and Set FStepoint
   VAR_TEMP   // added for the SCL form of the ladder/FBD networks
      _w1 : Bool;
   END_VAR
BEGIN

REGION Network 1
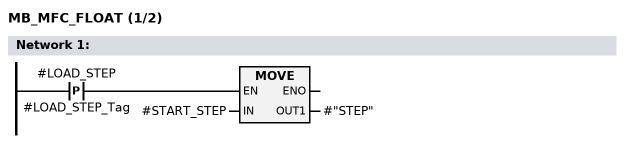
   RUNG wire#powerrail
      P_Contact(operand := #LOAD_STEP, bit := #LOAD_STEP_Tag)
      Move(in := #START_STEP, out1 => #"STEP")
   END_RUNG
   // the same network as SCL:
   #_w1 := #LOAD_STEP AND NOT #LOAD_STEP_Tag;   // rising edge of #LOAD_STEP
   #LOAD_STEP_Tag := #LOAD_STEP;
   IF #_w1 THEN #"STEP" := #START_STEP; END_IF;
END_REGION

REGION Network 2
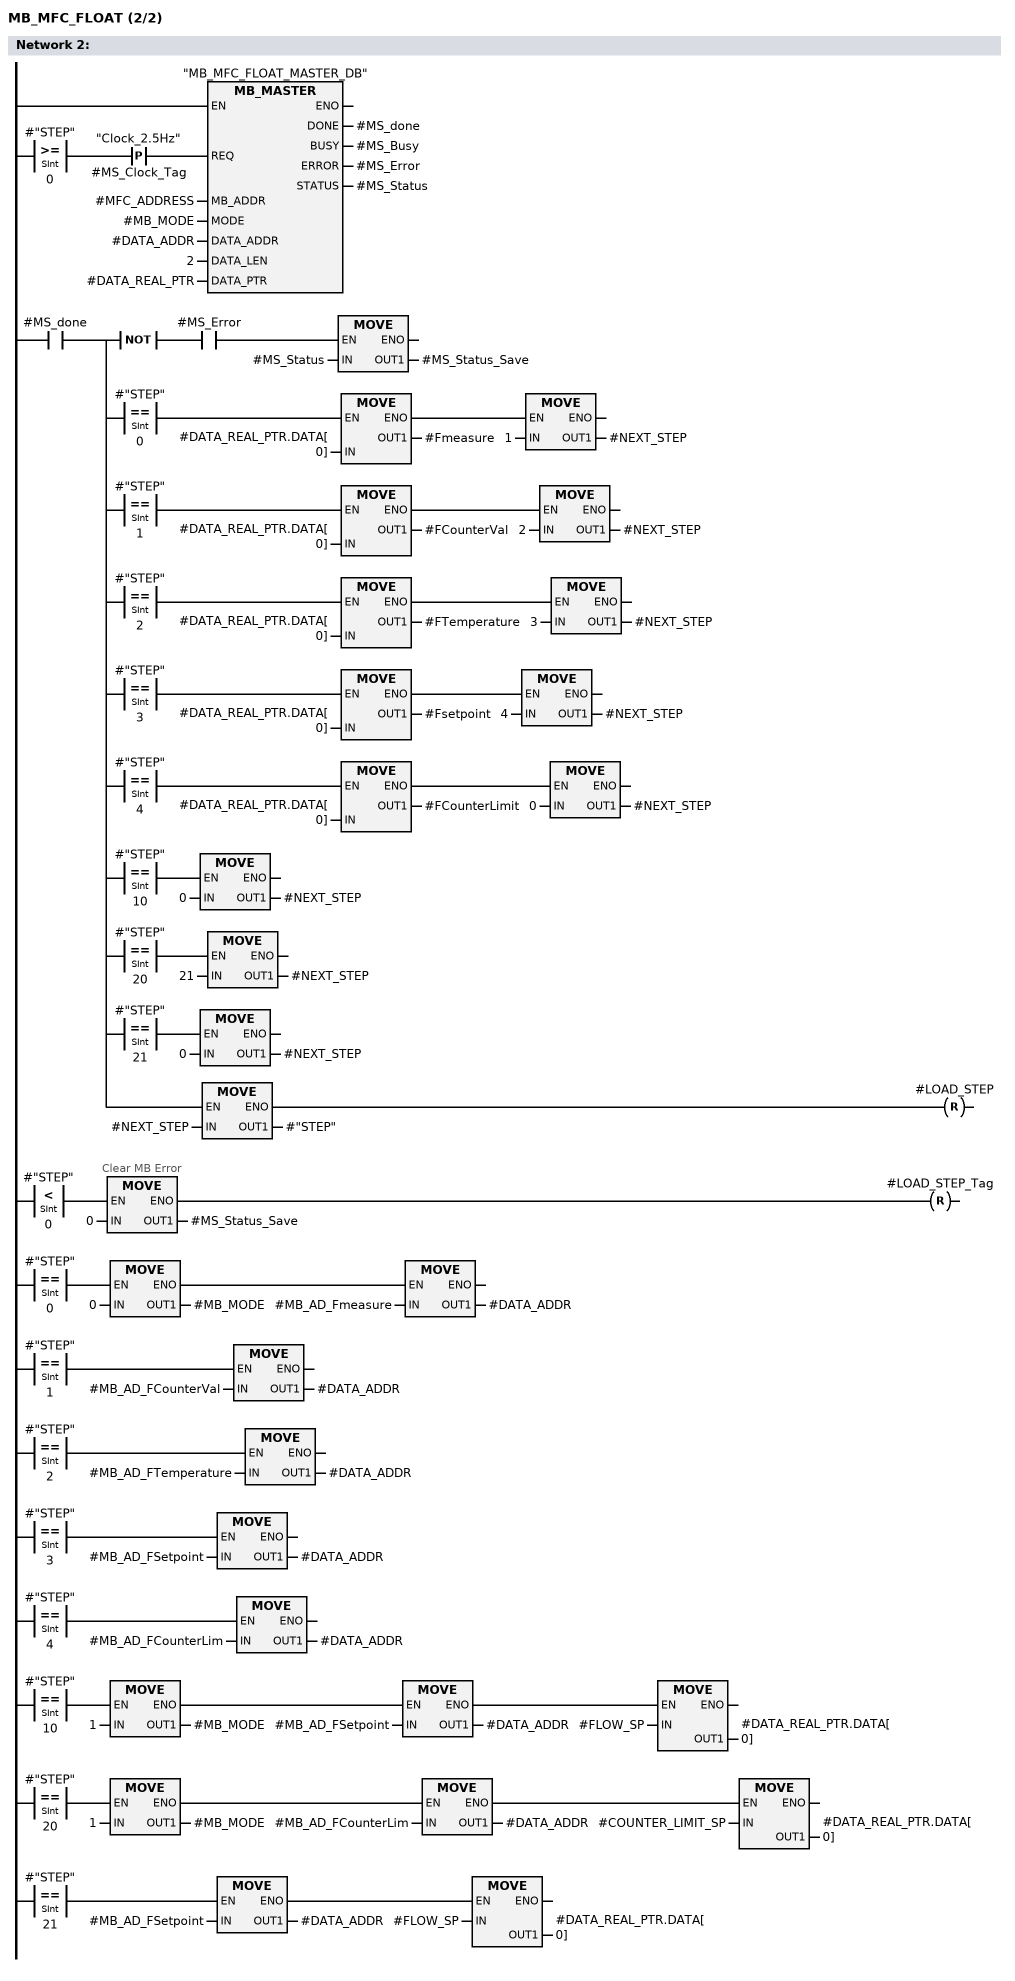
   #_w1 := (#"STEP" >= 0) AND "Clock_2.5Hz" AND NOT #MS_Clock_Tag;   // rising edge of "Clock_2.5Hz"
   #MS_Clock_Tag := "Clock_2.5Hz";
   "MB_MFC_FLOAT_MASTER_DB"(REQ := #_w1,   // MB_MASTER
                           MB_ADDR := #MFC_ADDRESS,
                           MODE := #MB_MODE,
                           DATA_ADDR := #DATA_ADDR,
                           DATA_LEN := 2,
                           DATA_PTR := #DATA_REAL_PTR,
                           DONE => #MS_done,
                           BUSY => #MS_Busy,
                           ERROR => #MS_Error,
                           STATUS => #MS_Status);
   IF NOT #MS_done AND #MS_Error THEN #MS_Status_Save := #MS_Status; END_IF;
   IF #MS_done AND (#"STEP" = 0) THEN
       #Fmeasure := #DATA_REAL_PTR.DATA[0];
       #NEXT_STEP := 1;
   END_IF;
   IF #MS_done AND (#"STEP" = 1) THEN
       #FCounterVal := #DATA_REAL_PTR.DATA[0];
       #NEXT_STEP := 2;
   END_IF;
   IF #MS_done AND (#"STEP" = 2) THEN
       #FTemperature := #DATA_REAL_PTR.DATA[0];
       #NEXT_STEP := 3;
   END_IF;
   IF #MS_done AND (#"STEP" = 3) THEN
       #Fsetpoint := #DATA_REAL_PTR.DATA[0];
       #NEXT_STEP := 4;
   END_IF;
   IF #MS_done AND (#"STEP" = 4) THEN
       #FCounterLimit := #DATA_REAL_PTR.DATA[0];
       #NEXT_STEP := 0;
   END_IF;
   IF #MS_done AND (#"STEP" = 10) THEN #NEXT_STEP := 0; END_IF;
   IF #MS_done AND (#"STEP" = 20) THEN #NEXT_STEP := 21; END_IF;
   IF #MS_done AND (#"STEP" = 21) THEN #NEXT_STEP := 0; END_IF;
   IF #MS_done THEN
       #"STEP" := #NEXT_STEP;
       #LOAD_STEP := FALSE;
   END_IF;
   IF #"STEP" < 0 THEN
       #MS_Status_Save := 0;   // Clear MB Error
       #LOAD_STEP_Tag := FALSE;
   END_IF;
   IF #"STEP" = 0 THEN
       #MB_MODE := 0;
       #DATA_ADDR := #MB_AD_Fmeasure;
   END_IF;
   IF #"STEP" = 1 THEN #DATA_ADDR := #MB_AD_FCounterVal; END_IF;
   IF #"STEP" = 2 THEN #DATA_ADDR := #MB_AD_FTemperature; END_IF;
   IF #"STEP" = 3 THEN #DATA_ADDR := #MB_AD_FSetpoint; END_IF;
   IF #"STEP" = 4 THEN #DATA_ADDR := #MB_AD_FCounterLim; END_IF;
   IF #"STEP" = 10 THEN
       #MB_MODE := 1;
       #DATA_ADDR := #MB_AD_FSetpoint;
       #DATA_REAL_PTR.DATA[0] := #FLOW_SP;
   END_IF;
   IF #"STEP" = 20 THEN
       #MB_MODE := 1;
       #DATA_ADDR := #MB_AD_FCounterLim;
       #DATA_REAL_PTR.DATA[0] := #COUNTER_LIMIT_SP;
   END_IF;
   IF #"STEP" = 21 THEN
       #DATA_ADDR := #MB_AD_FSetpoint;
       #DATA_REAL_PTR.DATA[0] := #FLOW_SP;
   END_IF;
END_REGION
END_FUNCTION_BLOCK

FUNCTION_BLOCK "MB_MFC_INT"   // FB2, LAD
{ S7_Optimized_Access := 'FALSE' }
VERSION : 0.1
// State Machine to control MFCs
// Steps 0-4: Measure Data
// Steps 10-12 Set Valve SP
// Steps 60: Set Control Mode
// Steps 68: Valve Fully Open (Purge)
// 
// Adresses: MFC201: 20 MFC601: 60
   VAR_TEMP   // added for the SCL form of the ladder/FBD networks
      _w1 : Bool;
   END_VAR
BEGIN

REGION Network 1
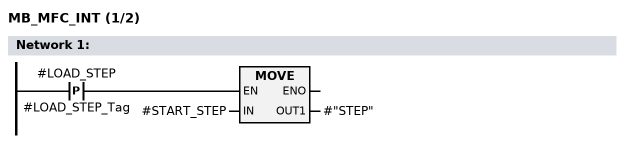
   RUNG wire#powerrail
      P_Contact(operand := #LOAD_STEP, bit := #LOAD_STEP_Tag)
      Move(in := #START_STEP, out1 => #"STEP")
   END_RUNG
   // the same network as SCL:
   #_w1 := #LOAD_STEP AND NOT #LOAD_STEP_Tag;   // rising edge of #LOAD_STEP
   #LOAD_STEP_Tag := #LOAD_STEP;
   IF #_w1 THEN #"STEP" := #START_STEP; END_IF;
END_REGION

REGION Network 2